   2553: 'Spare_Fault_2553', class No Acknowledgement, trigger "DB302_HMI_Faults_Carrier39_Faults_3" bit 8
   2554: 'Spare_Fault_2554', class No Acknowledgement, trigger "DB302_HMI_Faults_Carrier39_Faults_3" bit 9
   2555: 'Spare_Fault_2555', class No Acknowledgement, trigger "DB302_HMI_Faults_Carrier39_Faults_3" bit 10
   2556: 'Spare_Fault_2556', class No Acknowledgement, trigger "DB302_HMI_Faults_Carrier39_Faults_3" bit 11
   2557: 'Spare_Fault_2557', class No Acknowledgement, trigger "DB302_HMI_Faults_Carrier39_Faults_3" bit 12
   2558: 'Spare_Fault_2558', class No Acknowledgement, trigger "DB302_HMI_Faults_Carrier39_Faults_3" bit 13
   2559: 'Spare_Fault_2559', class No Acknowledgement, trigger "DB302_HMI_Faults_Carrier39_Faults_3" bit 14
   2560: 'Spare_Fault_2560', class No Acknowledgement, trigger "DB302_HMI_Faults_Carrier39_Faults_3" bit 15
   2561: 'Carrier 40 Disconnect Open Power Fault DI11.0', class No Acknowledgement, trigger "DB302_HMI_Faults_Carrier40_Faults_0" bit 0
   2562: 'Carrier 40 Drive Profinet Comm Fault', class No Acknowledgement, trigger "DB302_HMI_Faults_Carrier40_Faults_0" bit 1
   2563: 'Carrier 40 Production Stop Not Reset', class No Acknowledgement, trigger "DB302_HMI_Faults_Carrier40_Faults_0" bit 2
   2564: 'Carrier 40 CB02122 Tripped', class No Acknowledgement, trigger "DB302_HMI_Faults_Carrier40_Faults_0" bit 3
   2565: 'Carrier 40 CB02123 Tripped', class No Acknowledgement, trigger "DB302_HMI_Faults_Carrier40_Faults_0" bit 4
   2566: 'Carrier 40 AUX1 CB Tripped', class No Acknowledgement, trigger "DB302_HMI_Faults_Carrier40_Faults_0" bit 5
   2567: 'Carrier 40 AUX2 CB Tripped', class No Acknowledgement, trigger "DB302_HMI_Faults_Carrier40_Faults_0" bit 6
   2568: 'Carrier 40 PLC Not Communicating', class No Acknowledgement, trigger "DB302_HMI_Faults_Carrier40_Faults_0" bit 7
   2569: 'Carrier 40 Safe Input Card Fault', class No Acknowledgement, trigger "DB302_HMI_Faults_Carrier40_Faults_0" bit 8
   2570: 'Carrier 40 Safe Output Card Fault', class No Acknowledgement, trigger "DB302_HMI_Faults_Carrier40_Faults_0" bit 9
   2571: 'Carrier 40 Standard Input Card Fault', class No Acknowledgement, trigger "DB302_HMI_Faults_Carrier40_Faults_0" bit 10
   2572: 'Carrier 40 Standard Output Card Fault', class No Acknowledgement, trigger "DB302_HMI_Faults_Carrier40_Faults_0" bit 11
   2573: 'Carrier 40 Encoder Position Fault', class No Acknowledgement, trigger "DB302_HMI_Faults_Carrier40_Faults_0" bit 12
   2574: 'Carrier 40 Encoder Internal Error', class No Acknowledgement, trigger "DB302_HMI_Faults_Carrier40_Faults_0" bit 13
   2575: 'Carrier 40 Encoder Comm Fault', class No Acknowledgement, trigger "DB302_HMI_Faults_Carrier40_Faults_0" bit 14
   2576: 'Carrier 40 HMI Comm Fault', class No Acknowledgement, trigger "DB302_HMI_Faults_Carrier40_Faults_0" bit 15
   2577: 'Carrier 40 Crash Detection Fault', class No Acknowledgement, trigger "DB302_HMI_Faults_Carrier40_Faults_1" bit 0
   2578: 'Carrier 40 Carrier Number Invalid', class No Acknowledgement, trigger "DB302_HMI_Faults_Carrier40_Faults_1" bit 1
   2579: 'Carrier 40 Drive: PROFINET configuration error', class No Acknowledgement, trigger "DB302_HMI_Faults_Carrier40_Faults_1" bit 2
   2580: 'Carrier 40 Drive: Error internal communications', class No Acknowledgement, trigger "DB302_HMI_Faults_Carrier40_Faults_1" bit 3
   2581: 'Carrier 40 Drive: Motor overtemperature', class No Acknowledgement, trigger "DB302_HMI_Faults_Carrier40_Faults_1" bit 4
   2582: 'Carrier 40 Drive: Motor overcurrent', class No Acknowledgement, trigger "DB302_HMI_Faults_Carrier40_Faults_1" bit 5
   2583: 'Carrier 40 Drive: Infeed or power unit not ready', class No Acknowledgement, trigger "DB302_HMI_Faults_Carrier40_Faults_1" bit 6
   2584: 'Carrier 40 Drive: Short-circuit/ground fault detected', class No Acknowledgement, trigger "DB302_HMI_Faults_Carrier40_Faults_1" bit 7
   2585: 'Carrier 40 Drive: PROFINET Setpoint timeout', class No Acknowledgement, trigger "DB302_HMI_Faults_Carrier40_Faults_1" bit 8
   2586: 'Carrier 40 Power unit: Overcurrent', class No Acknowledgement, trigger "DB302_HMI_Faults_Carrier40_Faults_1" bit 9
   2587: 'Carrier 40 Power unit: DC link voltage overvoltage', class No Acknowledgement, trigger "DB302_HMI_Faults_Carrier40_Faults_1" bit 10
   2588: 'Carrier 40 Power unit: DC link voltage undervoltage', class No Acknowledgement, trigger "DB302_HMI_Faults_Carrier40_Faults_1" bit 11
   2589: 'Carrier 40 Power unit: Line phase failure in main circuit', class No Acknowledgement, trigger "DB302_HMI_Faults_Carrier40_Faults_1" bit 12
   2590: 'Carrier 40 Power unit: Phase failure motor cable', class No Acknowledgement, trigger "DB302_HMI_Faults_Carrier40_Faults_1" bit 13
   2591: 'Carrier 40 Power unit: Ground fault', class No Acknowledgement, trigger "DB302_HMI_Faults_Carrier40_Faults_1" bit 14
   2592: 'Spare_Fault_2592', class No Acknowledgement, trigger "DB302_HMI_Faults_Carrier40_Faults_1" bit 15
   2593: 'Carrier 40 Motion Off Fault', class No Acknowledgement, trigger "DB302_HMI_Faults_Carrier40_Faults_2" bit 0
   2594: 'Carrier 40 Motion On Fault', class No Acknowledgement, trigger "DB302_HMI_Faults_Carrier40_Faults_2" bit 1
   2595: 'Carrier 40 Spacing Fault', class No Acknowledgement, trigger "DB302_HMI_Faults_Carrier40_Faults_2" bit 2
   2596: 'Carrier 40 Duplicate Carrier Number Fault', class No Acknowledgement, trigger "DB302_HMI_Faults_Carrier40_Faults_2" bit 3
   2597: 'Spare_Fault_2597', class No Acknowledgement, trigger "DB302_HMI_Faults_Carrier40_Faults_2" bit 4
   2598: 'Spare_Fault_2598', class No Acknowledgement, trigger "DB302_HMI_Faults_Carrier40_Faults_2" bit 5
   2599: 'Spare_Fault_2599', class No Acknowledgement, trigger "DB302_HMI_Faults_Carrier40_Faults_2" bit 6
   2600: 'Spare_Fault_2600', class No Acknowledgement, trigger "DB302_HMI_Faults_Carrier40_Faults_2" bit 7
   2601: 'Spare_Fault_2601', class No Acknowledgement, trigger "DB302_HMI_Faults_Carrier40_Faults_2" bit 8
   2602: 'Spare_Fault_2602', class No Acknowledgement, trigger "DB302_HMI_Faults_Carrier40_Faults_2" bit 9
   2603: 'Spare_Fault_2603', class No Acknowledgement, trigger "DB302_HMI_Faults_Carrier40_Faults_2" bit 10
   2604: 'Spare_Fault_2604', class No Acknowledgement, trigger "DB302_HMI_Faults_Carrier40_Faults_2" bit 11
   2605: 'Spare_Fault_2605', class No Acknowledgement, trigger "DB302_HMI_Faults_Carrier40_Faults_2" bit 12
   2606: 'Spare_Fault_2606', class No Acknowledgement, trigger "DB302_HMI_Faults_Carrier40_Faults_2" bit 13
   2607: 'Spare_Fault_2607', class No Acknowledgement, trigger "DB302_HMI_Faults_Carrier40_Faults_2" bit 14
   2608: 'Spare_Fault_2608', class No Acknowledgement, trigger "DB302_HMI_Faults_Carrier40_Faults_2" bit 15
   2609: 'Spare_Fault_2609', class No Acknowledgement, trigger "DB302_HMI_Faults_Carrier40_Faults_3" bit 0
   2610: 'Spare_Fault_2610', class No Acknowledgement, trigger "DB302_HMI_Faults_Carrier40_Faults_3" bit 1
   2611: 'Spare_Fault_2611', class No Acknowledgement, trigger "DB302_HMI_Faults_Carrier40_Faults_3" bit 2
   2612: 'Spare_Fault_2612', class No Acknowledgement, trigger "DB302_HMI_Faults_Carrier40_Faults_3" bit 3
   2613: 'Spare_Fault_2613', class No Acknowledgement, trigger "DB302_HMI_Faults_Carrier40_Faults_3" bit 4
   2614: 'Spare_Fault_2614', class No Acknowledgement, trigger "DB302_HMI_Faults_Carrier40_Faults_3" bit 5
   2615: 'Spare_Fault_2615', class No Acknowledgement, trigger "DB302_HMI_Faults_Carrier40_Faults_3" bit 6
   2616: 'Spare_Fault_2616', class No Acknowledgement, trigger "DB302_HMI_Faults_Carrier40_Faults_3" bit 7
   2617: 'Spare_Fault_2617', class No Acknowledgement, trigger "DB302_HMI_Faults_Carrier40_Faults_3" bit 8
   2618: 'Spare_Fault_2618', class No Acknowledgement, trigger "DB302_HMI_Faults_Carrier40_Faults_3" bit 9
   2619: 'Spare_Fault_2619', class No Acknowledgement, trigger "DB302_HMI_Faults_Carrier40_Faults_3" bit 10
   2620: 'Spare_Fault_2620', class No Acknowledgement, trigger "DB302_HMI_Faults_Carrier40_Faults_3" bit 11
   2621: 'Spare_Fault_2621', class No Acknowledgement, trigger "DB302_HMI_Faults_Carrier40_Faults_3" bit 12
   2622: 'Spare_Fault_2622', class No Acknowledgement, trigger "DB302_HMI_Faults_Carrier40_Faults_3" bit 13
   2623: 'Spare_Fault_2623', class No Acknowledgement, trigger "DB302_HMI_Faults_Carrier40_Faults_3" bit 14
   2624: 'Spare_Fault_2624', class No Acknowledgement, trigger "DB302_HMI_Faults_Carrier40_Faults_3" bit 15
   2625: 'Carrier 41 Disconnect Open Power Fault DI11.0', class No Acknowledgement, trigger "DB302_HMI_Faults_Carrier41_Faults_0" bit 0
   2626: 'Carrier 41 Drive Profinet Comm Fault', class No Acknowledgement, trigger "DB302_HMI_Faults_Carrier41_Faults_0" bit 1
   2627: 'Carrier 41 Production Stop Not Reset', class No Acknowledgement, trigger "DB302_HMI_Faults_Carrier41_Faults_0" bit 2
   2628: 'Carrier 41 CB02122 Tripped', class No Acknowledgement, trigger "DB302_HMI_Faults_Carrier41_Faults_0" bit 3
   2629: 'Carrier 41 CB02123 Tripped', class No Acknowledgement, trigger "DB302_HMI_Faults_Carrier41_Faults_0" bit 4
   2630: 'Carrier 41 AUX1 CB Tripped', class No Acknowledgement, trigger "DB302_HMI_Faults_Carrier41_Faults_0" bit 5
   2631: 'Carrier 41 AUX2 CB Tripped', class No Acknowledgement, trigger "DB302_HMI_Faults_Carrier41_Faults_0" bit 6
   2632: 'Carrier 41 PLC Not Communicating', class No Acknowledgement, trigger "DB302_HMI_Faults_Carrier41_Faults_0" bit 7
   2633: 'Carrier 41 Safe Input Card Fault', class No Acknowledgement, trigger "DB302_HMI_Faults_Carrier41_Faults_0" bit 8
   2634: 'Carrier 41 Safe Output Card Fault', class No Acknowledgement, trigger "DB302_HMI_Faults_Carrier41_Faults_0" bit 9
   2635: 'Carrier 41 Standard Input Card Fault', class No Acknowledgement, trigger "DB302_HMI_Faults_Carrier41_Faults_0" bit 10
   2636: 'Carrier 41 Standard Output Card Fault', class No Acknowledgement, trigger "DB302_HMI_Faults_Carrier41_Faults_0" bit 11
   2637: 'Carrier 41 Encoder Position Fault', class No Acknowledgement, trigger "DB302_HMI_Faults_Carrier41_Faults_0" bit 12
   2638: 'Carrier 41 Encoder Internal Error', class No Acknowledgement, trigger "DB302_HMI_Faults_Carrier41_Faults_0" bit 13
   2639: 'Carrier 41 Encoder Comm Fault', class No Acknowledgement, trigger "DB302_HMI_Faults_Carrier41_Faults_0" bit 14
   2640: 'Carrier 41 HMI Comm Fault', class No Acknowledgement, trigger "DB302_HMI_Faults_Carrier41_Faults_0" bit 15
   2641: 'Carrier 41 Crash Detection Fault', class No Acknowledgement, trigger "DB302_HMI_Faults_Carrier41_Faults_1" bit 0
   2642: 'Carrier 41 Carrier Number Invalid', class No Acknowledgement, trigger "DB302_HMI_Faults_Carrier41_Faults_1" bit 1
   2643: 'Carrier 41 Drive: PROFINET configuration error', class No Acknowledgement, trigger "DB302_HMI_Faults_Carrier41_Faults_1" bit 2
   2644: 'Carrier 41 Drive: Error internal communications', class No Acknowledgement, trigger "DB302_HMI_Faults_Carrier41_Faults_1" bit 3
   2645: 'Carrier 41 Drive: Motor overtemperature', class No Acknowledgement, trigger "DB302_HMI_Faults_Carrier41_Faults_1" bit 4
   2646: 'Carrier 41 Drive: Motor overcurrent', class No Acknowledgement, trigger "DB302_HMI_Faults_Carrier41_Faults_1" bit 5
   2647: 'Carrier 41 Drive: Infeed or power unit not ready', class No Acknowledgement, trigger "DB302_HMI_Faults_Carrier41_Faults_1" bit 6
   2648: 'Carrier 41 Drive: Short-circuit/ground fault detected', class No Acknowledgement, trigger "DB302_HMI_Faults_Carrier41_Faults_1" bit 7
   2649: 'Carrier 41 Drive: PROFINET Setpoint timeout', class No Acknowledgement, trigger "DB302_HMI_Faults_Carrier41_Faults_1" bit 8
   2650: 'Carrier 41 Power unit: Overcurrent', class No Acknowledgement, trigger "DB302_HMI_Faults_Carrier41_Faults_1" bit 9
   2651: 'Carrier 41 Power unit: DC link voltage overvoltage', class No Acknowledgement, trigger "DB302_HMI_Faults_Carrier41_Faults_1" bit 10
   2652: 'Carrier 41 Power unit: DC link voltage undervoltage', class No Acknowledgement, trigger "DB302_HMI_Faults_Carrier41_Faults_1" bit 11
   2653: 'Carrier 41 Power unit: Line phase failure in main circuit', class No Acknowledgement, trigger "DB302_HMI_Faults_Carrier41_Faults_1" bit 12
   2654: 'Carrier 41 Power unit: Phase failure motor cable', class No Acknowledgement, trigger "DB302_HMI_Faults_Carrier41_Faults_1" bit 13
   2655: 'Carrier 41 Power unit: Ground fault', class No Acknowledgement, trigger "DB302_HMI_Faults_Carrier41_Faults_1" bit 14
   2656: 'Spare_Fault_2656', class No Acknowledgement, trigger "DB302_HMI_Faults_Carrier41_Faults_1" bit 15
   2657: 'Carrier 41 Motion Off Fault', class No Acknowledgement, trigger "DB302_HMI_Faults_Carrier41_Faults_2" bit 0
   2658: 'Carrier 41 Motion On Fault', class No Acknowledgement, trigger "DB302_HMI_Faults_Carrier41_Faults_2" bit 1
   2659: 'Carrier 41 Spacing Fault', class No Acknowledgement, trigger "DB302_HMI_Faults_Carrier41_Faults_2" bit 2
   2660: 'Carrier 41 Duplicate Carrier Number Fault', class No Acknowledgement, trigger "DB302_HMI_Faults_Carrier41_Faults_2" bit 3
   2661: 'Spare_Fault_2661', class No Acknowledgement, trigger "DB302_HMI_Faults_Carrier41_Faults_2" bit 4
   2662: 'Spare_Fault_2662', class No Acknowledgement, trigger "DB302_HMI_Faults_Carrier41_Faults_2" bit 5
   2663: 'Spare_Fault_2663', class No Acknowledgement, trigger "DB302_HMI_Faults_Carrier41_Faults_2" bit 6
   2664: 'Spare_Fault_2664', class No Acknowledgement, trigger "DB302_HMI_Faults_Carrier41_Faults_2" bit 7
   2665: 'Spare_Fault_2665', class No Acknowledgement, trigger "DB302_HMI_Faults_Carrier41_Faults_2" bit 8
   2666: 'Spare_Fault_2666', class No Acknowledgement, trigger "DB302_HMI_Faults_Carrier41_Faults_2" bit 9
   2667: 'Spare_Fault_2667', class No Acknowledgement, trigger "DB302_HMI_Faults_Carrier41_Faults_2" bit 10
   2668: 'Spare_Fault_2668', class No Acknowledgement, trigger "DB302_HMI_Faults_Carrier41_Faults_2" bit 11
   2669: 'Spare_Fault_2669', class No Acknowledgement, trigger "DB302_HMI_Faults_Carrier41_Faults_2" bit 12
   2670: 'Spare_Fault_2670', class No Acknowledgement, trigger "DB302_HMI_Faults_Carrier41_Faults_2" bit 13
   2671: 'Spare_Fault_2671', class No Acknowledgement, trigger "DB302_HMI_Faults_Carrier41_Faults_2" bit 14
   2672: 'Spare_Fault_2672', class No Acknowledgement, trigger "DB302_HMI_Faults_Carrier41_Faults_2" bit 15
   2673: 'Spare_Fault_2673', class No Acknowledgement, trigger "DB302_HMI_Faults_Carrier41_Faults_3" bit 0
   2674: 'Spare_Fault_2674', class No Acknowledgement, trigger "DB302_HMI_Faults_Carrier41_Faults_3" bit 1
   2675: 'Spare_Fault_2675', class No Acknowledgement, trigger "DB302_HMI_Faults_Carrier41_Faults_3" bit 2
   2676: 'Spare_Fault_2676', class No Acknowledgement, trigger "DB302_HMI_Faults_Carrier41_Faults_3" bit 3
   2677: 'Spare_Fault_2677', class No Acknowledgement, trigger "DB302_HMI_Faults_Carrier41_Faults_3" bit 4
   2678: 'Spare_Fault_2678', class No Acknowledgement, trigger "DB302_HMI_Faults_Carrier41_Faults_3" bit 5
   2679: 'Spare_Fault_2679', class No Acknowledgement, trigger "DB302_HMI_Faults_Carrier41_Faults_3" bit 6
   2680: 'Spare_Fault_2680', class No Acknowledgement, trigger "DB302_HMI_Faults_Carrier41_Faults_3" bit 7
   2681: 'Spare_Fault_2681', class No Acknowledgement, trigger "DB302_HMI_Faults_Carrier41_Faults_3" bit 8
   2682: 'Spare_Fault_2682', class No Acknowledgement, trigger "DB302_HMI_Faults_Carrier41_Faults_3" bit 9
   2683: 'Spare_Fault_2683', class No Acknowledgement, trigger "DB302_HMI_Faults_Carrier41_Faults_3" bit 10
   2684: 'Spare_Fault_2684', class No Acknowledgement, trigger "DB302_HMI_Faults_Carrier41_Faults_3" bit 11
   2685: 'Spare_Fault_2685', class No Acknowledgement, trigger "DB302_HMI_Faults_Carrier41_Faults_3" bit 12
   2686: 'Spare_Fault_2686', class No Acknowledgement, trigger "DB302_HMI_Faults_Carrier41_Faults_3" bit 13
   2687: 'Spare_Fault_2687', class No Acknowledgement, trigger "DB302_HMI_Faults_Carrier41_Faults_3" bit 14
   2688: 'Spare_Fault_2688', class No Acknowledgement, trigger "DB302_HMI_Faults_Carrier41_Faults_3" bit 15
   2689: 'Carrier 42 Disconnect Open Power Fault DI11.0', class No Acknowledgement, trigger "DB302_HMI_Faults_Carrier42_Faults_0" bit 0
   2690: 'Carrier 42 Drive Profinet Comm Fault', class No Acknowledgement, trigger "DB302_HMI_Faults_Carrier42_Faults_0" bit 1
   2691: 'Carrier 42 Production Stop Not Reset', class No Acknowledgement, trigger "DB302_HMI_Faults_Carrier42_Faults_0" bit 2
   2692: 'Carrier 42 CB02122 Tripped', class No Acknowledgement, trigger "DB302_HMI_Faults_Carrier42_Faults_0" bit 3
   2693: 'Carrier 42 CB02123 Tripped', class No Acknowledgement, trigger "DB302_HMI_Faults_Carrier42_Faults_0" bit 4
   2694: 'Carrier 42 AUX1 CB Tripped', class No Acknowledgement, trigger "DB302_HMI_Faults_Carrier42_Faults_0" bit 5
   2695: 'Carrier 42 AUX2 CB Tripped', class No Acknowledgement, trigger "DB302_HMI_Faults_Carrier42_Faults_0" bit 6
   2696: 'Carrier 42 PLC Not Communicating', class No Acknowledgement, trigger "DB302_HMI_Faults_Carrier42_Faults_0" bit 7
   2697: 'Carrier 42 Safe Input Card Fault', class No Acknowledgement, trigger "DB302_HMI_Faults_Carrier42_Faults_0" bit 8
   2698: 'Carrier 42 Safe Output Card Fault', class No Acknowledgement, trigger "DB302_HMI_Faults_Carrier42_Faults_0" bit 9
   2699: 'Carrier 42 Standard Input Card Fault', class No Acknowledgement, trigger "DB302_HMI_Faults_Carrier42_Faults_0" bit 10
   2700: 'Carrier 42 Standard Output Card Fault', class No Acknowledgement, trigger "DB302_HMI_Faults_Carrier42_Faults_0" bit 11
   2701: 'Carrier 42 Encoder Position Fault', class No Acknowledgement, trigger "DB302_HMI_Faults_Carrier42_Faults_0" bit 12
   2702: 'Carrier 42 Encoder Internal Error', class No Acknowledgement, trigger "DB302_HMI_Faults_Carrier42_Faults_0" bit 13
   2703: 'Carrier 42 Encoder Comm Fault', class No Acknowledgement, trigger "DB302_HMI_Faults_Carrier42_Faults_0" bit 14
   2704: 'Carrier 42 HMI Comm Fault', class No Acknowledgement, trigger "DB302_HMI_Faults_Carrier42_Faults_0" bit 15
   2705: 'Carrier 42 Crash Detection Fault', class No Acknowledgement, trigger "DB302_HMI_Faults_Carrier42_Faults_1" bit 0
   2706: 'Carrier 42 Carrier Number Invalid', class No Acknowledgement, trigger "DB302_HMI_Faults_Carrier42_Faults_1" bit 1
   2707: 'Carrier 42 Drive: PROFINET configuration error', class No Acknowledgement, trigger "DB302_HMI_Faults_Carrier42_Faults_1" bit 2
   2708: 'Carrier 42 Drive: Error internal communications', class No Acknowledgement, trigger "DB302_HMI_Faults_Carrier42_Faults_1" bit 3
   2709: 'Carrier 42 Drive: Motor overtemperature', class No Acknowledgement, trigger "DB302_HMI_Faults_Carrier42_Faults_1" bit 4
   2710: 'Carrier 42 Drive: Motor overcurrent', class No Acknowledgement, trigger "DB302_HMI_Faults_Carrier42_Faults_1" bit 5
   2711: 'Carrier 42 Drive: Infeed or power unit not ready', class No Acknowledgement, trigger "DB302_HMI_Faults_Carrier42_Faults_1" bit 6
   2712: 'Carrier 42 Drive: Short-circuit/ground fault detected', class No Acknowledgement, trigger "DB302_HMI_Faults_Carrier42_Faults_1" bit 7
   2713: 'Carrier 42 Drive: PROFINET Setpoint timeout', class No Acknowledgement, trigger "DB302_HMI_Faults_Carrier42_Faults_1" bit 8
   2714: 'Carrier 42 Power unit: Overcurrent', class No Acknowledgement, trigger "DB302_HMI_Faults_Carrier42_Faults_1" bit 9
   2715: 'Carrier 42 Power unit: DC link voltage overvoltage', class No Acknowledgement, trigger "DB302_HMI_Faults_Carrier42_Faults_1" bit 10
   2716: 'Carrier 42 Power unit: DC link voltage undervoltage', class No Acknowledgement, trigger "DB302_HMI_Faults_Carrier42_Faults_1" bit 11
   2717: 'Carrier 42 Power unit: Line phase failure in main circuit', class No Acknowledgement, trigger "DB302_HMI_Faults_Carrier42_Faults_1" bit 12
   2718: 'Carrier 42 Power unit: Phase failure motor cable', class No Acknowledgement, trigger "DB302_HMI_Faults_Carrier42_Faults_1" bit 13
   2719: 'Carrier 42 Power unit: Ground fault', class No Acknowledgement, trigger "DB302_HMI_Faults_Carrier42_Faults_1" bit 14
   2720: 'Spare_Fault_2720', class No Acknowledgement, trigger "DB302_HMI_Faults_Carrier42_Faults_1" bit 15
   2721: 'Carrier 42 Motion Off Fault', class No Acknowledgement, trigger "DB302_HMI_Faults_Carrier42_Faults_2" bit 0
   2722: 'Carrier 42 Motion On Fault', class No Acknowledgement, trigger "DB302_HMI_Faults_Carrier42_Faults_2" bit 1
   2723: 'Carrier 42 Spacing Fault', class No Acknowledgement, trigger "DB302_HMI_Faults_Carrier42_Faults_2" bit 2
   2724: 'Carrier 42 Duplicate Carrier Number Fault', class No Acknowledgement, trigger "DB302_HMI_Faults_Carrier42_Faults_2" bit 3
   2725: 'Spare_Fault_2725', class No Acknowledgement, trigger "DB302_HMI_Faults_Carrier42_Faults_2" bit 4
   2726: 'Spare_Fault_2726', class No Acknowledgement, trigger "DB302_HMI_Faults_Carrier42_Faults_2" bit 5
   2727: 'Spare_Fault_2727', class No Acknowledgement, trigger "DB302_HMI_Faults_Carrier42_Faults_2" bit 6
   2728: 'Spare_Fault_2728', class No Acknowledgement, trigger "DB302_HMI_Faults_Carrier42_Faults_2" bit 7
   2729: 'Spare_Fault_2729', class No Acknowledgement, trigger "DB302_HMI_Faults_Carrier42_Faults_2" bit 8
   2730: 'Spare_Fault_2730', class No Acknowledgement, trigger "DB302_HMI_Faults_Carrier42_Faults_2" bit 9
   2731: 'Spare_Fault_2731', class No Acknowledgement, trigger "DB302_HMI_Faults_Carrier42_Faults_2" bit 10
   2732: 'Spare_Fault_2732', class No Acknowledgement, trigger "DB302_HMI_Faults_Carrier42_Faults_2" bit 11
   2733: 'Spare_Fault_2733', class No Acknowledgement, trigger "DB302_HMI_Faults_Carrier42_Faults_2" bit 12
   2734: 'Spare_Fault_2734', class No Acknowledgement, trigger "DB302_HMI_Faults_Carrier42_Faults_2" bit 13
   2735: 'Spare_Fault_2735', class No Acknowledgement, trigger "DB302_HMI_Faults_Carrier42_Faults_2" bit 14
   2736: 'Spare_Fault_2736', class No Acknowledgement, trigger "DB302_HMI_Faults_Carrier42_Faults_2" bit 15
   2737: 'Spare_Fault_2737', class No Acknowledgement, trigger "DB302_HMI_Faults_Carrier42_Faults_3" bit 0
   2738: 'Spare_Fault_2738', class No Acknowledgement, trigger "DB302_HMI_Faults_Carrier42_Faults_3" bit 1
   2739: 'Spare_Fault_2739', class No Acknowledgement, trigger "DB302_HMI_Faults_Carrier42_Faults_3" bit 2
   2740: 'Spare_Fault_2740', class No Acknowledgement, trigger "DB302_HMI_Faults_Carrier42_Faults_3" bit 3
   2741: 'Spare_Fault_2741', class No Acknowledgement, trigger "DB302_HMI_Faults_Carrier42_Faults_3" bit 4
   2742: 'Spare_Fault_2742', class No Acknowledgement, trigger "DB302_HMI_Faults_Carrier42_Faults_3" bit 5
   2743: 'Spare_Fault_2743', class No Acknowledgement, trigger "DB302_HMI_Faults_Carrier42_Faults_3" bit 6
   2744: 'Spare_Fault_2744', class No Acknowledgement, trigger "DB302_HMI_Faults_Carrier42_Faults_3" bit 7
   2745: 'Spare_Fault_2745', class No Acknowledgement, trigger "DB302_HMI_Faults_Carrier42_Faults_3" bit 8
   2746: 'Spare_Fault_2746', class No Acknowledgement, trigger "DB302_HMI_Faults_Carrier42_Faults_3" bit 9
   2747: 'Spare_Fault_2747', class No Acknowledgement, trigger "DB302_HMI_Faults_Carrier42_Faults_3" bit 10
   2748: 'Spare_Fault_2748', class No Acknowledgement, trigger "DB302_HMI_Faults_Carrier42_Faults_3" bit 11
   2749: 'Spare_Fault_2749', class No Acknowledgement, trigger "DB302_HMI_Faults_Carrier42_Faults_3" bit 12
   2750: 'Spare_Fault_2750', class No Acknowledgement, trigger "DB302_HMI_Faults_Carrier42_Faults_3" bit 13
   2751: 'Spare_Fault_2751', class No Acknowledgement, trigger "DB302_HMI_Faults_Carrier42_Faults_3" bit 14
   2752: 'Spare_Fault_2752', class No Acknowledgement, trigger "DB302_HMI_Faults_Carrier42_Faults_3" bit 15
   2753: 'Carrier 43 Disconnect Open Power Fault DI11.0', class No Acknowledgement, trigger "DB302_HMI_Faults_Carrier43_Faults_0" bit 0
   2754: 'Carrier 43 Drive Profinet Comm Fault', class No Acknowledgement, trigger "DB302_HMI_Faults_Carrier43_Faults_0" bit 1
   2755: 'Carrier 43 Production Stop Not Reset', class No Acknowledgement, trigger "DB302_HMI_Faults_Carrier43_Faults_0" bit 2
   2756: 'Carrier 43 CB02122 Tripped', class No Acknowledgement, trigger "DB302_HMI_Faults_Carrier43_Faults_0" bit 3
   2757: 'Carrier 43 CB02123 Tripped', class No Acknowledgement, trigger "DB302_HMI_Faults_Carrier43_Faults_0" bit 4
   2758: 'Carrier 43 AUX1 CB Tripped', class No Acknowledgement, trigger "DB302_HMI_Faults_Carrier43_Faults_0" bit 5
   2759: 'Carrier 43 AUX2 CB Tripped', class No Acknowledgement, trigger "DB302_HMI_Faults_Carrier43_Faults_0" bit 6
   2760: 'Carrier 43 PLC Not Communicating', class No Acknowledgement, trigger "DB302_HMI_Faults_Carrier43_Faults_0" bit 7
   2761: 'Carrier 43 Safe Input Card Fault', class No Acknowledgement, trigger "DB302_HMI_Faults_Carrier43_Faults_0" bit 8
   2762: 'Carrier 43 Safe Output Card Fault', class No Acknowledgement, trigger "DB302_HMI_Faults_Carrier43_Faults_0" bit 9
   2763: 'Carrier 43 Standard Input Card Fault', class No Acknowledgement, trigger "DB302_HMI_Faults_Carrier43_Faults_0" bit 10
   2764: 'Carrier 43 Standard Output Card Fault', class No Acknowledgement, trigger "DB302_HMI_Faults_Carrier43_Faults_0" bit 11
   2765: 'Carrier 43 Encoder Position Fault', class No Acknowledgement, trigger "DB302_HMI_Faults_Carrier43_Faults_0" bit 12
   2766: 'Carrier 43 Encoder Internal Error', class No Acknowledgement, trigger "DB302_HMI_Faults_Carrier43_Faults_0" bit 13
   2767: 'Carrier 43 Encoder Comm Fault', class No Acknowledgement, trigger "DB302_HMI_Faults_Carrier43_Faults_0" bit 14
   2768: 'Carrier 43 HMI Comm Fault', class No Acknowledgement, trigger "DB302_HMI_Faults_Carrier43_Faults_0" bit 15
   2769: 'Carrier 43 Crash Detection Fault', class No Acknowledgement, trigger "DB302_HMI_Faults_Carrier43_Faults_1" bit 0
   2770: 'Carrier 43 Carrier Number Invalid', class No Acknowledgement, trigger "DB302_HMI_Faults_Carrier43_Faults_1" bit 1
   2771: 'Carrier 43 Drive: PROFINET configuration error', class No Acknowledgement, trigger "DB302_HMI_Faults_Carrier43_Faults_1" bit 2
   2772: 'Carrier 43 Drive: Error internal communications', class No Acknowledgement, trigger "DB302_HMI_Faults_Carrier43_Faults_1" bit 3
   2773: 'Carrier 43 Drive: Motor overtemperature', class No Acknowledgement, trigger "DB302_HMI_Faults_Carrier43_Faults_1" bit 4
   2774: 'Carrier 43 Drive: Motor overcurrent', class No Acknowledgement, trigger "DB302_HMI_Faults_Carrier43_Faults_1" bit 5
   2775: 'Carrier 43 Drive: Infeed or power unit not ready', class No Acknowledgement, trigger "DB302_HMI_Faults_Carrier43_Faults_1" bit 6
   2776: 'Carrier 43 Drive: Short-circuit/ground fault detected', class No Acknowledgement, trigger "DB302_HMI_Faults_Carrier43_Faults_1" bit 7
   2777: 'Carrier 43 Drive: PROFINET Setpoint timeout', class No Acknowledgement, trigger "DB302_HMI_Faults_Carrier43_Faults_1" bit 8
   2778: 'Carrier 43 Power unit: Overcurrent', class No Acknowledgement, trigger "DB302_HMI_Faults_Carrier43_Faults_1" bit 9
   2779: 'Carrier 43 Power unit: DC link voltage overvoltage', class No Acknowledgement, trigger "DB302_HMI_Faults_Carrier43_Faults_1" bit 10
   2780: 'Carrier 43 Power unit: DC link voltage undervoltage', class No Acknowledgement, trigger "DB302_HMI_Faults_Carrier43_Faults_1" bit 11
   2781: 'Carrier 43 Power unit: Line phase failure in main circuit', class No Acknowledgement, trigger "DB302_HMI_Faults_Carrier43_Faults_1" bit 12
   2782: 'Carrier 43 Power unit: Phase failure motor cable', class No Acknowledgement, trigger "DB302_HMI_Faults_Carrier43_Faults_1" bit 13
   2783: 'Carrier 43 Power unit: Ground fault', class No Acknowledgement, trigger "DB302_HMI_Faults_Carrier43_Faults_1" bit 14
   2784: 'Spare_Fault_2784', class No Acknowledgement, trigger "DB302_HMI_Faults_Carrier43_Faults_1" bit 15
   2785: 'Carrier 43 Motion Off Fault', class No Acknowledgement, trigger "DB302_HMI_Faults_Carrier43_Faults_2" bit 0
   2786: 'Carrier 43 Motion On Fault', class No Acknowledgement, trigger "DB302_HMI_Faults_Carrier43_Faults_2" bit 1
   2787: 'Carrier 43 Spacing Fault', class No Acknowledgement, trigger "DB302_HMI_Faults_Carrier43_Faults_2" bit 2
   2788: 'Carrier 43 Duplicate Carrier Number Fault', class No Acknowledgement, trigger "DB302_HMI_Faults_Carrier43_Faults_2" bit 3
   2789: 'Spare_Fault_2789', class No Acknowledgement, trigger "DB302_HMI_Faults_Carrier43_Faults_2" bit 4
   2790: 'Spare_Fault_2790', class No Acknowledgement, trigger "DB302_HMI_Faults_Carrier43_Faults_2" bit 5
   2791: 'Spare_Fault_2791', class No Acknowledgement, trigger "DB302_HMI_Faults_Carrier43_Faults_2" bit 6
   2792: 'Spare_Fault_2792', class No Acknowledgement, trigger "DB302_HMI_Faults_Carrier43_Faults_2" bit 7
   2793: 'Spare_Fault_2793', class No Acknowledgement, trigger "DB302_HMI_Faults_Carrier43_Faults_2" bit 8
   2794: 'Spare_Fault_2794', class No Acknowledgement, trigger "DB302_HMI_Faults_Carrier43_Faults_2" bit 9
   2795: 'Spare_Fault_2795', class No Acknowledgement, trigger "DB302_HMI_Faults_Carrier43_Faults_2" bit 10
   2796: 'Spare_Fault_2796', class No Acknowledgement, trigger "DB302_HMI_Faults_Carrier43_Faults_2" bit 11
   2797: 'Spare_Fault_2797', class No Acknowledgement, trigger "DB302_HMI_Faults_Carrier43_Faults_2" bit 12
   2798: 'Spare_Fault_2798', class No Acknowledgement, trigger "DB302_HMI_Faults_Carrier43_Faults_2" bit 13
   2799: 'Spare_Fault_2799', class No Acknowledgement, trigger "DB302_HMI_Faults_Carrier43_Faults_2" bit 14
   2800: 'Spare_Fault_2800', class No Acknowledgement, trigger "DB302_HMI_Faults_Carrier43_Faults_2" bit 15
   2801: 'Spare_Fault_2801', class No Acknowledgement, trigger "DB302_HMI_Faults_Carrier43_Faults_3" bit 0
   2802: 'Spare_Fault_2802', class No Acknowledgement, trigger "DB302_HMI_Faults_Carrier43_Faults_3" bit 1
   2803: 'Spare_Fault_2803', class No Acknowledgement, trigger "DB302_HMI_Faults_Carrier43_Faults_3" bit 2
   2804: 'Spare_Fault_2804', class No Acknowledgement, trigger "DB302_HMI_Faults_Carrier43_Faults_3" bit 3
   2805: 'Spare_Fault_2805', class No Acknowledgement, trigger "DB302_HMI_Faults_Carrier43_Faults_3" bit 4
   2806: 'Spare_Fault_2806', class No Acknowledgement, trigger "DB302_HMI_Faults_Carrier43_Faults_3" bit 5
   2807: 'Spare_Fault_2807', class No Acknowledgement, trigger "DB302_HMI_Faults_Carrier43_Faults_3" bit 6
   2808: 'Spare_Fault_2808', class No Acknowledgement, trigger "DB302_HMI_Faults_Carrier43_Faults_3" bit 7
   2809: 'Spare_Fault_2809', class No Acknowledgement, trigger "DB302_HMI_Faults_Carrier43_Faults_3" bit 8
   2810: 'Spare_Fault_2810', class No Acknowledgement, trigger "DB302_HMI_Faults_Carrier43_Faults_3" bit 9
   2811: 'Spare_Fault_2811', class No Acknowledgement, trigger "DB302_HMI_Faults_Carrier43_Faults_3" bit 10
   2812: 'Spare_Fault_2812', class No Acknowledgement, trigger "DB302_HMI_Faults_Carrier43_Faults_3" bit 11
   2813: 'Spare_Fault_2813', class No Acknowledgement, trigger "DB302_HMI_Faults_Carrier43_Faults_3" bit 12
   2814: 'Spare_Fault_2814', class No Acknowledgement, trigger "DB302_HMI_Faults_Carrier43_Faults_3" bit 13
   2815: 'Spare_Fault_2815', class No Acknowledgement, trigger "DB302_HMI_Faults_Carrier43_Faults_3" bit 14
   2816: 'Spare_Fault_2816', class No Acknowledgement, trigger "DB302_HMI_Faults_Carrier43_Faults_3" bit 15
   2817: 'Carrier 44 Disconnect Open Power Fault DI11.0', class No Acknowledgement, trigger "DB302_HMI_Faults_Carrier44_Faults_0" bit 0
   2818: 'Carrier 44 Drive Profinet Comm Fault', class No Acknowledgement, trigger "DB302_HMI_Faults_Carrier44_Faults_0" bit 1
   2819: 'Carrier 44 Production Stop Not Reset', class No Acknowledgement, trigger "DB302_HMI_Faults_Carrier44_Faults_0" bit 2
   2820: 'Carrier 44 CB02122 Tripped', class No Acknowledgement, trigger "DB302_HMI_Faults_Carrier44_Faults_0" bit 3
   2821: 'Carrier 44 CB02123 Tripped', class No Acknowledgement, trigger "DB302_HMI_Faults_Carrier44_Faults_0" bit 4
   2822: 'Carrier 44 AUX1 CB Tripped', class No Acknowledgement, trigger "DB302_HMI_Faults_Carrier44_Faults_0" bit 5
   2823: 'Carrier 44 AUX2 CB Tripped', class No Acknowledgement, trigger "DB302_HMI_Faults_Carrier44_Faults_0" bit 6
   2824: 'Carrier 44 PLC Not Communicating', class No Acknowledgement, trigger "DB302_HMI_Faults_Carrier44_Faults_0" bit 7
   2825: 'Carrier 44 Safe Input Card Fault', class No Acknowledgement, trigger "DB302_HMI_Faults_Carrier44_Faults_0" bit 8
   2826: 'Carrier 44 Safe Output Card Fault', class No Acknowledgement, trigger "DB302_HMI_Faults_Carrier44_Faults_0" bit 9
   2827: 'Carrier 44 Standard Input Card Fault', class No Acknowledgement, trigger "DB302_HMI_Faults_Carrier44_Faults_0" bit 10
   2828: 'Carrier 44 Standard Output Card Fault', class No Acknowledgement, trigger "DB302_HMI_Faults_Carrier44_Faults_0" bit 11
   2829: 'Carrier 44 Encoder Position Fault', class No Acknowledgement, trigger "DB302_HMI_Faults_Carrier44_Faults_0" bit 12
   2830: 'Carrier 44 Encoder Internal Error', class No Acknowledgement, trigger "DB302_HMI_Faults_Carrier44_Faults_0" bit 13
   2831: 'Carrier 44 Encoder Comm Fault', class No Acknowledgement, trigger "DB302_HMI_Faults_Carrier44_Faults_0" bit 14
   2832: 'Carrier 44 HMI Comm Fault', class No Acknowledgement, trigger "DB302_HMI_Faults_Carrier44_Faults_0" bit 15
   2833: 'Carrier 44 Crash Detection Fault', class No Acknowledgement, trigger "DB302_HMI_Faults_Carrier44_Faults_1" bit 0
   2834: 'Carrier 44 Carrier Number Invalid', class No Acknowledgement, trigger "DB302_HMI_Faults_Carrier44_Faults_1" bit 1
   2835: 'Carrier 44 Drive: PROFINET configuration error', class No Acknowledgement, trigger "DB302_HMI_Faults_Carrier44_Faults_1" bit 2
   2836: 'Carrier 44 Drive: Error internal communications', class No Acknowledgement, trigger "DB302_HMI_Faults_Carrier44_Faults_1" bit 3
   2837: 'Carrier 44 Drive: Motor overtemperature', class No Acknowledgement, trigger "DB302_HMI_Faults_Carrier44_Faults_1" bit 4
   2838: 'Carrier 44 Drive: Motor overcurrent', class No Acknowledgement, trigger "DB302_HMI_Faults_Carrier44_Faults_1" bit 5
   2839: 'Carrier 44 Drive: Infeed or power unit not ready', class No Acknowledgement, trigger "DB302_HMI_Faults_Carrier44_Faults_1" bit 6
   2840: 'Carrier 44 Drive: Short-circuit/ground fault detected', class No Acknowledgement, trigger "DB302_HMI_Faults_Carrier44_Faults_1" bit 7
   2841: 'Carrier 44 Drive: PROFINET Setpoint timeout', class No Acknowledgement, trigger "DB302_HMI_Faults_Carrier44_Faults_1" bit 8
   2842: 'Carrier 44 Power unit: Overcurrent', class No Acknowledgement, trigger "DB302_HMI_Faults_Carrier44_Faults_1" bit 9
   2843: 'Carrier 44 Power unit: DC link voltage overvoltage', class No Acknowledgement, trigger "DB302_HMI_Faults_Carrier44_Faults_1" bit 10
   2844: 'Carrier 44 Power unit: DC link voltage undervoltage', class No Acknowledgement, trigger "DB302_HMI_Faults_Carrier44_Faults_1" bit 11
   2845: 'Carrier 44 Power unit: Line phase failure in main circuit', class No Acknowledgement, trigger "DB302_HMI_Faults_Carrier44_Faults_1" bit 12
   2846: 'Carrier 44 Power unit: Phase failure motor cable', class No Acknowledgement, trigger "DB302_HMI_Faults_Carrier44_Faults_1" bit 13
   2847: 'Carrier 44 Power unit: Ground fault', class No Acknowledgement, trigger "DB302_HMI_Faults_Carrier44_Faults_1" bit 14
   2848: 'Spare_Fault_2848', class No Acknowledgement, trigger "DB302_HMI_Faults_Carrier44_Faults_1" bit 15
   2849: 'Carrier 44 Motion Off Fault', class No Acknowledgement, trigger "DB302_HMI_Faults_Carrier44_Faults_2" bit 0
   2850: 'Carrier 44 Motion On Fault', class No Acknowledgement, trigger "DB302_HMI_Faults_Carrier44_Faults_2" bit 1
   2851: 'Carrier 44 Spacing Fault', class No Acknowledgement, trigger "DB302_HMI_Faults_Carrier44_Faults_2" bit 2
   2852: 'Carrier 44 Duplicate Carrier Number Fault', class No Acknowledgement, trigger "DB302_HMI_Faults_Carrier44_Faults_2" bit 3
   2853: 'Spare_Fault_2853', class No Acknowledgement, trigger "DB302_HMI_Faults_Carrier44_Faults_2" bit 4
   2854: 'Spare_Fault_2854', class No Acknowledgement, trigger "DB302_HMI_Faults_Carrier44_Faults_2" bit 5
   2855: 'Spare_Fault_2855', class No Acknowledgement, trigger "DB302_HMI_Faults_Carrier44_Faults_2" bit 6
   2856: 'Spare_Fault_2856', class No Acknowledgement, trigger "DB302_HMI_Faults_Carrier44_Faults_2" bit 7
   2857: 'Spare_Fault_2857', class No Acknowledgement, trigger "DB302_HMI_Faults_Carrier44_Faults_2" bit 8
   2858: 'Spare_Fault_2858', class No Acknowledgement, trigger "DB302_HMI_Faults_Carrier44_Faults_2" bit 9
   2859: 'Spare_Fault_2859', class No Acknowledgement, trigger "DB302_HMI_Faults_Carrier44_Faults_2" bit 10
   2860: 'Spare_Fault_2860', class No Acknowledgement, trigger "DB302_HMI_Faults_Carrier44_Faults_2" bit 11
   2861: 'Spare_Fault_2861', class No Acknowledgement, trigger "DB302_HMI_Faults_Carrier44_Faults_2" bit 12
   2862: 'Spare_Fault_2862', class No Acknowledgement, trigger "DB302_HMI_Faults_Carrier44_Faults_2" bit 13
   2863: 'Spare_Fault_2863', class No Acknowledgement, trigger "DB302_HMI_Faults_Carrier44_Faults_2" bit 14
   2864: 'Spare_Fault_2864', class No Acknowledgement, trigger "DB302_HMI_Faults_Carrier44_Faults_2" bit 15
   2865: 'Spare_Fault_2865', class No Acknowledgement, trigger "DB302_HMI_Faults_Carrier44_Faults_3" bit 0
   2866: 'Spare_Fault_2866', class No Acknowledgement, trigger "DB302_HMI_Faults_Carrier44_Faults_3" bit 1
   2867: 'Spare_Fault_2867', class No Acknowledgement, trigger "DB302_HMI_Faults_Carrier44_Faults_3" bit 2
   2868: 'Spare_Fault_2868', class No Acknowledgement, trigger "DB302_HMI_Faults_Carrier44_Faults_3" bit 3
   2869: 'Spare_Fault_2869', class No Acknowledgement, trigger "DB302_HMI_Faults_Carrier44_Faults_3" bit 4
   2870: 'Spare_Fault_2870', class No Acknowledgement, trigger "DB302_HMI_Faults_Carrier44_Faults_3" bit 5
   2871: 'Spare_Fault_2871', class No Acknowledgement, trigger "DB302_HMI_Faults_Carrier44_Faults_3" bit 6
   2872: 'Spare_Fault_2872', class No Acknowledgement, trigger "DB302_HMI_Faults_Carrier44_Faults_3" bit 7
   2873: 'Spare_Fault_2873', class No Acknowledgement, trigger "DB302_HMI_Faults_Carrier44_Faults_3" bit 8
   2874: 'Spare_Fault_2874', class No Acknowledgement, trigger "DB302_HMI_Faults_Carrier44_Faults_3" bit 9
   2875: 'Spare_Fault_2875', class No Acknowledgement, trigger "DB302_HMI_Faults_Carrier44_Faults_3" bit 10
   2876: 'Spare_Fault_2876', class No Acknowledgement, trigger "DB302_HMI_Faults_Carrier44_Faults_3" bit 11
   2877: 'Spare_Fault_2877', class No Acknowledgement, trigger "DB302_HMI_Faults_Carrier44_Faults_3" bit 12
   2878: 'Spare_Fault_2878', class No Acknowledgement, trigger "DB302_HMI_Faults_Carrier44_Faults_3" bit 13
   2879: 'Spare_Fault_2879', class No Acknowledgement, trigger "DB302_HMI_Faults_Carrier44_Faults_3" bit 14
   2880: 'Spare_Fault_2880', class No Acknowledgement, trigger "DB302_HMI_Faults_Carrier44_Faults_3" bit 15
   2881: 'Carrier 45 Disconnect Open Power Fault DI11.0', class No Acknowledgement, trigger "DB302_HMI_Faults_Carrier45_Faults_0" bit 0
   2882: 'Carrier 45 Drive Profinet Comm Fault', class No Acknowledgement, trigger "DB302_HMI_Faults_Carrier45_Faults_0" bit 1
   2883: 'Carrier 45 Production Stop Not Reset', class No Acknowledgement, trigger "DB302_HMI_Faults_Carrier45_Faults_0" bit 2
   2884: 'Carrier 45 CB02122 Tripped', class No Acknowledgement, trigger "DB302_HMI_Faults_Carrier45_Faults_0" bit 3
   2885: 'Carrier 45 CB02123 Tripped', class No Acknowledgement, trigger "DB302_HMI_Faults_Carrier45_Faults_0" bit 4
   2886: 'Carrier 45 AUX1 CB Tripped', class No Acknowledgement, trigger "DB302_HMI_Faults_Carrier45_Faults_0" bit 5
   2887: 'Carrier 45 AUX2 CB Tripped', class No Acknowledgement, trigger "DB302_HMI_Faults_Carrier45_Faults_0" bit 6
   2888: 'Carrier 45 PLC Not Communicating', class No Acknowledgement, trigger "DB302_HMI_Faults_Carrier45_Faults_0" bit 7
   2889: 'Carrier 45 Safe Input Card Fault', class No Acknowledgement, trigger "DB302_HMI_Faults_Carrier45_Faults_0" bit 8
   2890: 'Carrier 45 Safe Output Card Fault', class No Acknowledgement, trigger "DB302_HMI_Faults_Carrier45_Faults_0" bit 9
   2891: 'Carrier 45 Standard Input Card Fault', class No Acknowledgement, trigger "DB302_HMI_Faults_Carrier45_Faults_0" bit 10
   2892: 'Carrier 45 Standard Output Card Fault', class No Acknowledgement, trigger "DB302_HMI_Faults_Carrier45_Faults_0" bit 11
   2893: 'Carrier 45 Encoder Position Fault', class No Acknowledgement, trigger "DB302_HMI_Faults_Carrier45_Faults_0" bit 12
   2894: 'Carrier 45 Encoder Internal Error', class No Acknowledgement, trigger "DB302_HMI_Faults_Carrier45_Faults_0" bit 13
   2895: 'Carrier 45 Encoder Comm Fault', class No Acknowledgement, trigger "DB302_HMI_Faults_Carrier45_Faults_0" bit 14
   2896: 'Carrier 45 HMI Comm Fault', class No Acknowledgement, trigger "DB302_HMI_Faults_Carrier45_Faults_0" bit 15
   2897: 'Carrier 45 Crash Detection Fault', class No Acknowledgement, trigger "DB302_HMI_Faults_Carrier45_Faults_1" bit 0
   2898: 'Carrier 45 Carrier Number Invalid', class No Acknowledgement, trigger "DB302_HMI_Faults_Carrier45_Faults_1" bit 1
   2899: 'Carrier 45 Drive: PROFINET configuration error', class No Acknowledgement, trigger "DB302_HMI_Faults_Carrier45_Faults_1" bit 2
   2900: 'Carrier 45 Drive: Error internal communications', class No Acknowledgement, trigger "DB302_HMI_Faults_Carrier45_Faults_1" bit 3
   2901: 'Carrier 45 Drive: Motor overtemperature', class No Acknowledgement, trigger "DB302_HMI_Faults_Carrier45_Faults_1" bit 4
   2902: 'Carrier 45 Drive: Motor overcurrent', class No Acknowledgement, trigger "DB302_HMI_Faults_Carrier45_Faults_1" bit 5
   2903: 'Carrier 45 Drive: Infeed or power unit not ready', class No Acknowledgement, trigger "DB302_HMI_Faults_Carrier45_Faults_1" bit 6
   2904: 'Carrier 45 Drive: Short-circuit/ground fault detected', class No Acknowledgement, trigger "DB302_HMI_Faults_Carrier45_Faults_1" bit 7
   2905: 'Carrier 45 Drive: PROFINET Setpoint timeout', class No Acknowledgement, trigger "DB302_HMI_Faults_Carrier45_Faults_1" bit 8
   2906: 'Carrier 45 Power unit: Overcurrent', class No Acknowledgement, trigger "DB302_HMI_Faults_Carrier45_Faults_1" bit 9
   2907: 'Carrier 45 Power unit: DC link voltage overvoltage', class No Acknowledgement, trigger "DB302_HMI_Faults_Carrier45_Faults_1" bit 10
   2908: 'Carrier 45 Power unit: DC link voltage undervoltage', class No Acknowledgement, trigger "DB302_HMI_Faults_Carrier45_Faults_1" bit 11
   2909: 'Carrier 45 Power unit: Line phase failure in main circuit', class No Acknowledgement, trigger "DB302_HMI_Faults_Carrier45_Faults_1" bit 12
   2910: 'Carrier 45 Power unit: Phase failure motor cable', class No Acknowledgement, trigger "DB302_HMI_Faults_Carrier45_Faults_1" bit 13
   2911: 'Carrier 45 Power unit: Ground fault', class No Acknowledgement, trigger "DB302_HMI_Faults_Carrier45_Faults_1" bit 14
   2912: 'Spare_Fault_2912', class No Acknowledgement, trigger "DB302_HMI_Faults_Carrier45_Faults_1" bit 15
   2913: 'Carrier 45 Motion Off Fault', class No Acknowledgement, trigger "DB302_HMI_Faults_Carrier45_Faults_2" bit 0
   2914: 'Carrier 45 Motion On Fault', class No Acknowledgement, trigger "DB302_HMI_Faults_Carrier45_Faults_2" bit 1
   2915: 'Carrier 45 Spacing Fault', class No Acknowledgement, trigger "DB302_HMI_Faults_Carrier45_Faults_2" bit 2
   2916: 'Carrier 45 Duplicate Carrier Number Fault', class No Acknowledgement, trigger "DB302_HMI_Faults_Carrier45_Faults_2" bit 3
   2917: 'Spare_Fault_2917', class No Acknowledgement, trigger "DB302_HMI_Faults_Carrier45_Faults_2" bit 4
   2918: 'Spare_Fault_2918', class No Acknowledgement, trigger "DB302_HMI_Faults_Carrier45_Faults_2" bit 5
   2919: 'Spare_Fault_2919', class No Acknowledgement, trigger "DB302_HMI_Faults_Carrier45_Faults_2" bit 6
   2920: 'Spare_Fault_2920', class No Acknowledgement, trigger "DB302_HMI_Faults_Carrier45_Faults_2" bit 7
   2921: 'Spare_Fault_2921', class No Acknowledgement, trigger "DB302_HMI_Faults_Carrier45_Faults_2" bit 8
   2922: 'Spare_Fault_2922', class No Acknowledgement, trigger "DB302_HMI_Faults_Carrier45_Faults_2" bit 9
   2923: 'Spare_Fault_2923', class No Acknowledgement, trigger "DB302_HMI_Faults_Carrier45_Faults_2" bit 10
   2924: 'Spare_Fault_2924', class No Acknowledgement, trigger "DB302_HMI_Faults_Carrier45_Faults_2" bit 11
   2925: 'Spare_Fault_2925', class No Acknowledgement, trigger "DB302_HMI_Faults_Carrier45_Faults_2" bit 12
   2926: 'Spare_Fault_2926', class No Acknowledgement, trigger "DB302_HMI_Faults_Carrier45_Faults_2" bit 13
   2927: 'Spare_Fault_2927', class No Acknowledgement, trigger "DB302_HMI_Faults_Carrier45_Faults_2" bit 14
   2928: 'Spare_Fault_2928', class No Acknowledgement, trigger "DB302_HMI_Faults_Carrier45_Faults_2" bit 15
   2929: 'Spare_Fault_2929', class No Acknowledgement, trigger "DB302_HMI_Faults_Carrier45_Faults_3" bit 0
   2930: 'Spare_Fault_2930', class No Acknowledgement, trigger "DB302_HMI_Faults_Carrier45_Faults_3" bit 1
   2931: 'Spare_Fault_2931', class No Acknowledgement, trigger "DB302_HMI_Faults_Carrier45_Faults_3" bit 2
   2932: 'Spare_Fault_2932', class No Acknowledgement, trigger "DB302_HMI_Faults_Carrier45_Faults_3" bit 3
   2933: 'Spare_Fault_2933', class No Acknowledgement, trigger "DB302_HMI_Faults_Carrier45_Faults_3" bit 4
   2934: 'Spare_Fault_2934', class No Acknowledgement, trigger "DB302_HMI_Faults_Carrier45_Faults_3" bit 5
   2935: 'Spare_Fault_2935', class No Acknowledgement, trigger "DB302_HMI_Faults_Carrier45_Faults_3" bit 6
   2936: 'Spare_Fault_2936', class No Acknowledgement, trigger "DB302_HMI_Faults_Carrier45_Faults_3" bit 7
   2937: 'Spare_Fault_2937', class No Acknowledgement, trigger "DB302_HMI_Faults_Carrier45_Faults_3" bit 8
   2938: 'Spare_Fault_2938', class No Acknowledgement, trigger "DB302_HMI_Faults_Carrier45_Faults_3" bit 9
   2939: 'Spare_Fault_2939', class No Acknowledgement, trigger "DB302_HMI_Faults_Carrier45_Faults_3" bit 10
   2940: 'Spare_Fault_2940', class No Acknowledgement, trigger "DB302_HMI_Faults_Carrier45_Faults_3" bit 11
   2941: 'Spare_Fault_2941', class No Acknowledgement, trigger "DB302_HMI_Faults_Carrier45_Faults_3" bit 12
   2942: 'Spare_Fault_2942', class No Acknowledgement, trigger "DB302_HMI_Faults_Carrier45_Faults_3" bit 13
   2943: 'Spare_Fault_2943', class No Acknowledgement, trigger "DB302_HMI_Faults_Carrier45_Faults_3" bit 14
   2944: 'Spare_Fault_2944', class No Acknowledgement, trigger "DB302_HMI_Faults_Carrier45_Faults_3" bit 15
   2945: 'Carrier 46 Disconnect Open Power Fault DI11.0', class No Acknowledgement, trigger "DB302_HMI_Faults_Carrier46_Faults_0" bit 0
   2946: 'Carrier 46 Drive Profinet Comm Fault', class No Acknowledgement, trigger "DB302_HMI_Faults_Carrier46_Faults_0" bit 1
   2947: 'Carrier 46 Production Stop Not Reset', class No Acknowledgement, trigger "DB302_HMI_Faults_Carrier46_Faults_0" bit 2
   2948: 'Carrier 46 CB02122 Tripped', class No Acknowledgement, trigger "DB302_HMI_Faults_Carrier46_Faults_0" bit 3
   2949: 'Carrier 46 CB02123 Tripped', class No Acknowledgement, trigger "DB302_HMI_Faults_Carrier46_Faults_0" bit 4
   2950: 'Carrier 46 AUX1 CB Tripped', class No Acknowledgement, trigger "DB302_HMI_Faults_Carrier46_Faults_0" bit 5
   2951: 'Carrier 46 AUX2 CB Tripped', class No Acknowledgement, trigger "DB302_HMI_Faults_Carrier46_Faults_0" bit 6
   2952: 'Carrier 46 PLC Not Communicating', class No Acknowledgement, trigger "DB302_HMI_Faults_Carrier46_Faults_0" bit 7
   2953: 'Carrier 46 Safe Input Card Fault', class No Acknowledgement, trigger "DB302_HMI_Faults_Carrier46_Faults_0" bit 8
   2954: 'Carrier 46 Safe Output Card Fault', class No Acknowledgement, trigger "DB302_HMI_Faults_Carrier46_Faults_0" bit 9
   2955: 'Carrier 46 Standard Input Card Fault', class No Acknowledgement, trigger "DB302_HMI_Faults_Carrier46_Faults_0" bit 10
   2956: 'Carrier 46 Standard Output Card Fault', class No Acknowledgement, trigger "DB302_HMI_Faults_Carrier46_Faults_0" bit 11
   2957: 'Carrier 46 Encoder Position Fault', class No Acknowledgement, trigger "DB302_HMI_Faults_Carrier46_Faults_0" bit 12
   2958: 'Carrier 46 Encoder Internal Error', class No Acknowledgement, trigger "DB302_HMI_Faults_Carrier46_Faults_0" bit 13
   2959: 'Carrier 46 Encoder Comm Fault', class No Acknowledgement, trigger "DB302_HMI_Faults_Carrier46_Faults_0" bit 14
   2960: 'Carrier 46 HMI Comm Fault', class No Acknowledgement, trigger "DB302_HMI_Faults_Carrier46_Faults_0" bit 15
   2961: 'Carrier 46 Crash Detection Fault', class No Acknowledgement, trigger "DB302_HMI_Faults_Carrier46_Faults_1" bit 0
   2962: 'Carrier 46 Carrier Number Invalid', class No Acknowledgement, trigger "DB302_HMI_Faults_Carrier46_Faults_1" bit 1
   2963: 'Carrier 46 Drive: PROFINET configuration error', class No Acknowledgement, trigger "DB302_HMI_Faults_Carrier46_Faults_1" bit 2
   2964: 'Carrier 46 Drive: Error internal communications', class No Acknowledgement, trigger "DB302_HMI_Faults_Carrier46_Faults_1" bit 3
   2965: 'Carrier 46 Drive: Motor overtemperature', class No Acknowledgement, trigger "DB302_HMI_Faults_Carrier46_Faults_1" bit 4
   2966: 'Carrier 46 Drive: Motor overcurrent', class No Acknowledgement, trigger "DB302_HMI_Faults_Carrier46_Faults_1" bit 5
   2967: 'Carrier 46 Drive: Infeed or power unit not ready', class No Acknowledgement, trigger "DB302_HMI_Faults_Carrier46_Faults_1" bit 6
   2968: 'Carrier 46 Drive: Short-circuit/ground fault detected', class No Acknowledgement, trigger "DB302_HMI_Faults_Carrier46_Faults_1" bit 7
   2969: 'Carrier 46 Drive: PROFINET Setpoint timeout', class No Acknowledgement, trigger "DB302_HMI_Faults_Carrier46_Faults_1" bit 8
   2970: 'Carrier 46 Power unit: Overcurrent', class No Acknowledgement, trigger "DB302_HMI_Faults_Carrier46_Faults_1" bit 9
   2971: 'Carrier 46 Power unit: DC link voltage overvoltage', class No Acknowledgement, trigger "DB302_HMI_Faults_Carrier46_Faults_1" bit 10
   2972: 'Carrier 46 Power unit: DC link voltage undervoltage', class No Acknowledgement, trigger "DB302_HMI_Faults_Carrier46_Faults_1" bit 11